REGION Network 14
   RUNG wire#powerrail
      "FC_ANIM_MOTOR"(Input_1 := "MP012-CO", Input_3 := "DB90".Static_6, Input_4 := "MP012-TO", Input_5 := "DB34".Static_24, Output_0 => "DB46".Static_2, Input_0 := wire#w1, Input_2 := wire#w2)
   END_RUNG
   RUNG wire#powerrail
      Contact( "MP012-Marcha" )
      I_Contact( "PRESOSTATO-TORRES" )
   END_RUNG wire#w1
   RUNG wire#powerrail
      Contact( "DB90".Static_110 )
      I_Contact( "DB90".Static_136 )
   END_RUNG wire#w2
   // the same network as SCL:
   "FC_ANIM_MOTOR"(Input_0 := "MP012-Marcha" AND NOT "PRESOSTATO-TORRES",
                   Input_1 := "MP012-CO",
                   Input_2 := "DB90".Static_110 AND NOT "DB90".Static_136,
                   Input_3 := "DB90".Static_6,
                   Input_4 := "MP012-TO",
                   Input_5 := "DB34".Static_24,
                   Output_0 => "DB46".Static_2);
END_REGION

REGION Network 15
   RUNG wire#powerrail
      "FC_ANIM_MOTOR"(Input_1 := "MP013-CO", Input_3 := "DB90".Static_7, Input_4 := "MP013-TO", Input_5 := "DB34".Static_26, Output_0 => "DB46".Static_3, Input_0 := wire#w1, Input_2 := wire#w2)
   END_RUNG
   RUNG wire#powerrail
      Contact( "MP013-Marcha" )
      I_Contact( "PRESOSTATO-TORRES" )
   END_RUNG wire#w1
   RUNG wire#powerrail
      Contact( "DB90".Static_111 )
      I_Contact( "DB90".Static_137 )
   END_RUNG wire#w2
   // the same network as SCL:
   "FC_ANIM_MOTOR"(Input_0 := "MP013-Marcha" AND NOT "PRESOSTATO-TORRES",
                   Input_1 := "MP013-CO",
                   Input_2 := "DB90".Static_111 AND NOT "DB90".Static_137,
                   Input_3 := "DB90".Static_7,
                   Input_4 := "MP013-TO",
                   Input_5 := "DB34".Static_26,
                   Output_0 => "DB46".Static_3);
END_REGION

REGION Network 16
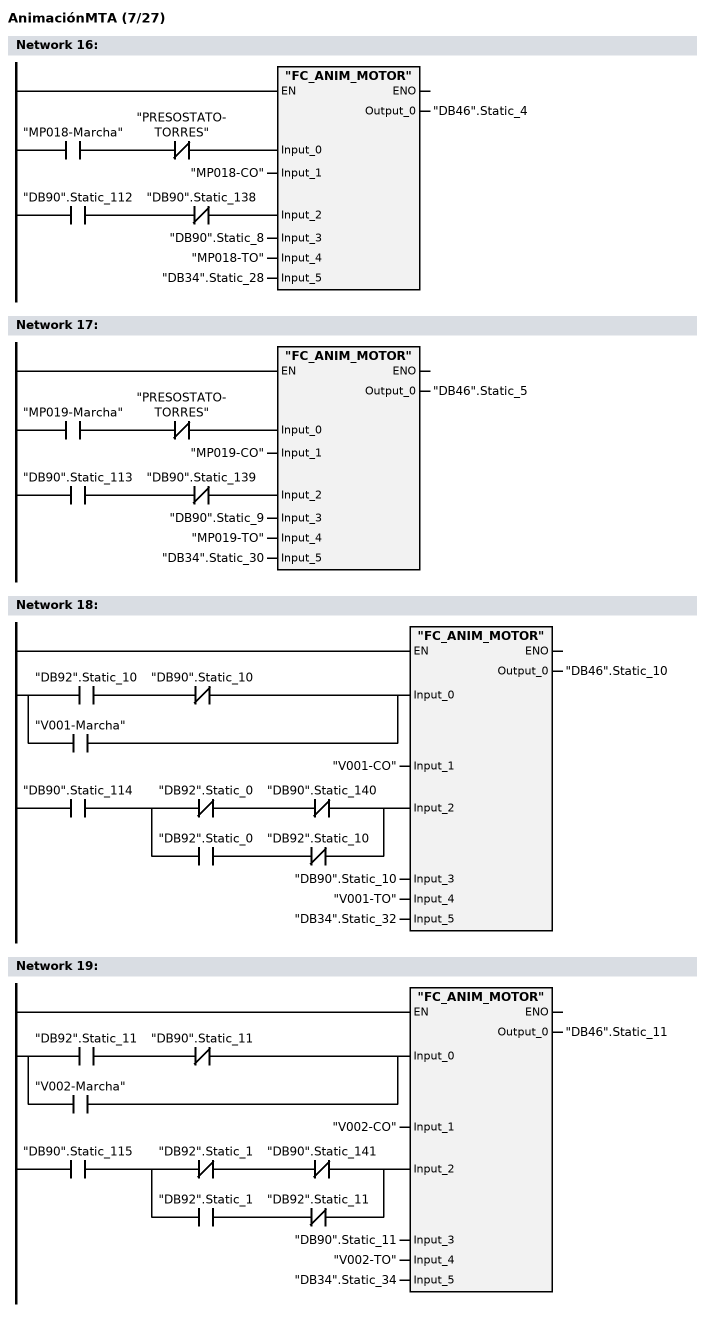
   RUNG wire#powerrail
      "FC_ANIM_MOTOR"(Input_1 := "MP018-CO", Input_3 := "DB90".Static_8, Input_4 := "MP018-TO", Input_5 := "DB34".Static_28, Output_0 => "DB46".Static_4, Input_0 := wire#w1, Input_2 := wire#w2)
   END_RUNG
   RUNG wire#powerrail
      Contact( "MP018-Marcha" )
      I_Contact( "PRESOSTATO-TORRES" )
   END_RUNG wire#w1
   RUNG wire#powerrail
      Contact( "DB90".Static_112 )
      I_Contact( "DB90".Static_138 )
   END_RUNG wire#w2
   // the same network as SCL:
   "FC_ANIM_MOTOR"(Input_0 := "MP018-Marcha" AND NOT "PRESOSTATO-TORRES",
                   Input_1 := "MP018-CO",
                   Input_2 := "DB90".Static_112 AND NOT "DB90".Static_138,
                   Input_3 := "DB90".Static_8,
                   Input_4 := "MP018-TO",
                   Input_5 := "DB34".Static_28,
                   Output_0 => "DB46".Static_4);
END_REGION

REGION Network 17
   RUNG wire#powerrail
      "FC_ANIM_MOTOR"(Input_1 := "MP019-CO", Input_3 := "DB90".Static_9, Input_4 := "MP019-TO", Input_5 := "DB34".Static_30, Output_0 => "DB46".Static_5, Input_0 := wire#w1, Input_2 := wire#w2)
   END_RUNG
   RUNG wire#powerrail
      Contact( "MP019-Marcha" )
      I_Contact( "PRESOSTATO-TORRES" )
   END_RUNG wire#w1
   RUNG wire#powerrail
      Contact( "DB90".Static_113 )
      I_Contact( "DB90".Static_139 )
   END_RUNG wire#w2
   // the same network as SCL:
   "FC_ANIM_MOTOR"(Input_0 := "MP019-Marcha" AND NOT "PRESOSTATO-TORRES",
                   Input_1 := "MP019-CO",
                   Input_2 := "DB90".Static_113 AND NOT "DB90".Static_139,
                   Input_3 := "DB90".Static_9,
                   Input_4 := "MP019-TO",
                   Input_5 := "DB34".Static_30,
                   Output_0 => "DB46".Static_5);
END_REGION

REGION Network 18
   "FC_ANIM_MOTOR"(Input_0 := "V001-Marcha" OR ("DB92".Static_10 AND NOT "DB90".Static_10),
                   Input_1 := "V001-CO",
                   Input_2 := "DB90".Static_114 AND ((NOT "DB92".Static_0 AND NOT "DB90".Static_140) OR ("DB92".Static_0 AND NOT "DB92".Static_10)),
                   Input_3 := "DB90".Static_10,
                   Input_4 := "V001-TO",
                   Input_5 := "DB34".Static_32,
                   Output_0 => "DB46".Static_10);
END_REGION

REGION Network 19
   "FC_ANIM_MOTOR"(Input_0 := "V002-Marcha" OR ("DB92".Static_11 AND NOT "DB90".Static_11),
                   Input_1 := "V002-CO",
                   Input_2 := "DB90".Static_115 AND ((NOT "DB92".Static_1 AND NOT "DB90".Static_141) OR ("DB92".Static_1 AND NOT "DB92".Static_11)),
                   Input_3 := "DB90".Static_11,
                   Input_4 := "V002-TO",
                   Input_5 := "DB34".Static_34,
                   Output_0 => "DB46".Static_11);
END_REGION

REGION Network 20
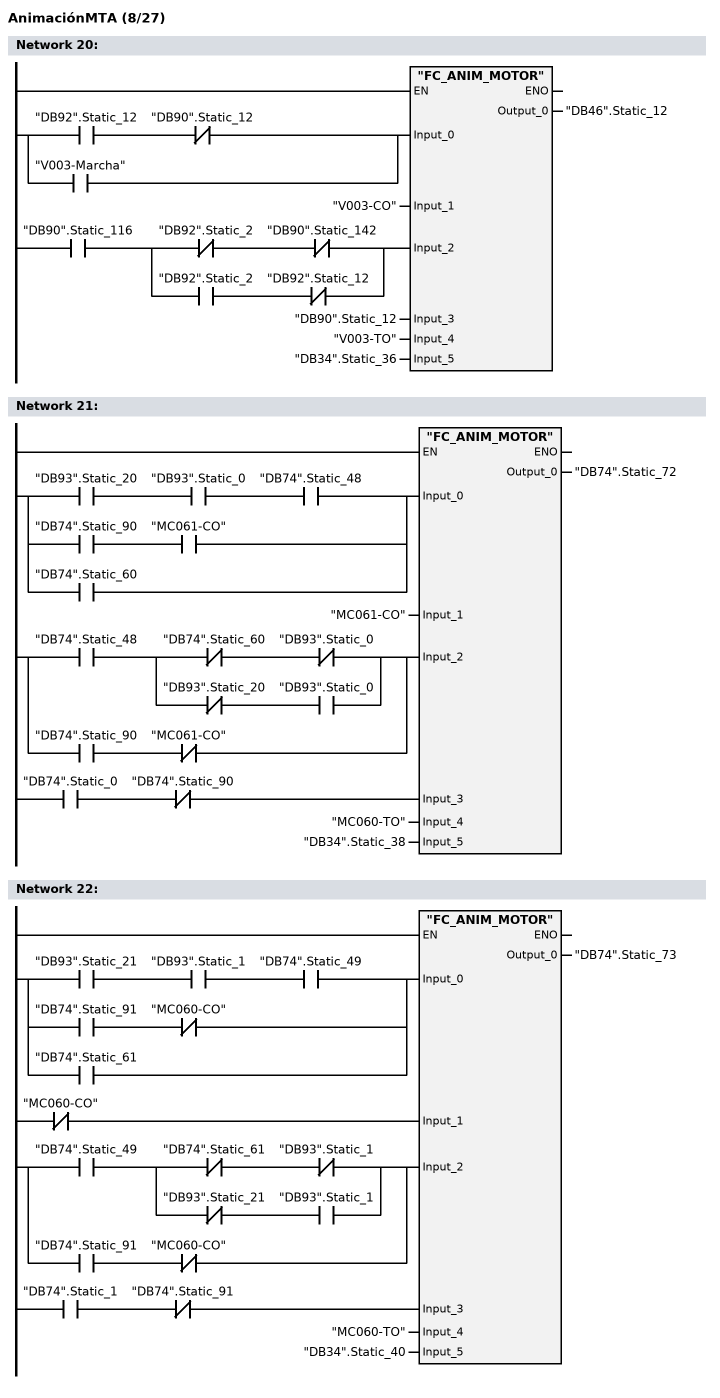
   "FC_ANIM_MOTOR"(Input_0 := "V003-Marcha" OR ("DB92".Static_12 AND NOT "DB90".Static_12),
                   Input_1 := "V003-CO",
                   Input_2 := "DB90".Static_116 AND ((NOT "DB92".Static_2 AND NOT "DB90".Static_142) OR ("DB92".Static_2 AND NOT "DB92".Static_12)),
                   Input_3 := "DB90".Static_12,
                   Input_4 := "V003-TO",
                   Input_5 := "DB34".Static_36,
                   Output_0 => "DB46".Static_12);
END_REGION

REGION Network 21
   "FC_ANIM_MOTOR"(Input_0 := "DB74".Static_60 OR ("DB93".Static_20 AND "DB93".Static_0 AND "DB74".Static_48) OR ("DB74".Static_90 AND "MC061-CO"),
                   Input_1 := "MC061-CO",
                   Input_2 := ("DB74".Static_48 AND ((NOT "DB74".Static_60 AND NOT "DB93".Static_0) OR (NOT "DB93".Static_20 AND "DB93".Static_0))) OR ("DB74".Static_90 AND NOT "MC061-CO"),
                   Input_3 := "DB74".Static_0 AND NOT "DB74".Static_90,
                   Input_4 := "MC060-TO",
                   Input_5 := "DB34".Static_38,
                   Output_0 => "DB74".Static_72);
END_REGION

REGION Network 22
   "FC_ANIM_MOTOR"(Input_0 := "DB74".Static_61 OR ("DB93".Static_21 AND "DB93".Static_1 AND "DB74".Static_49) OR ("DB74".Static_91 AND NOT "MC060-CO"),
                   Input_1 := NOT "MC060-CO",
                   Input_2 := ("DB74".Static_49 AND ((NOT "DB74".Static_61 AND NOT "DB93".Static_1) OR (NOT "DB93".Static_21 AND "DB93".Static_1))) OR ("DB74".Static_91 AND NOT "MC060-CO"),
                   Input_3 := "DB74".Static_1 AND NOT "DB74".Static_91,
                   Input_4 := "MC060-TO",
                   Input_5 := "DB34".Static_40,
                   Output_0 => "DB74".Static_73);
END_REGION

REGION Network 23
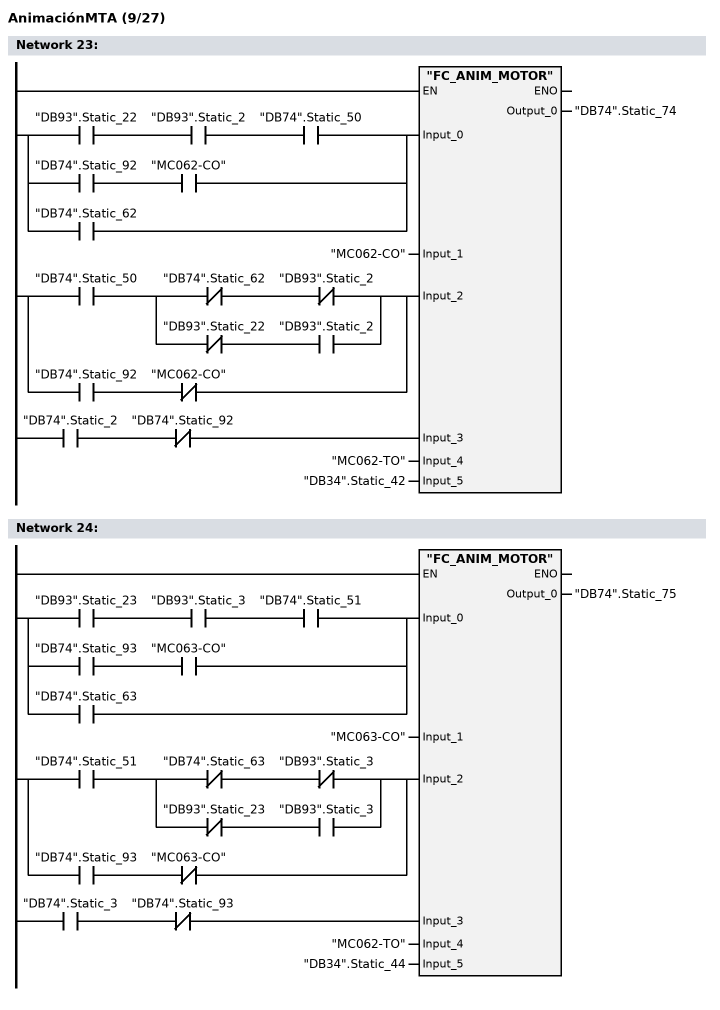
   "FC_ANIM_MOTOR"(Input_0 := "DB74".Static_62 OR ("DB93".Static_22 AND "DB93".Static_2 AND "DB74".Static_50) OR ("DB74".Static_92 AND "MC062-CO"),
                   Input_1 := "MC062-CO",
                   Input_2 := ("DB74".Static_50 AND ((NOT "DB74".Static_62 AND NOT "DB93".Static_2) OR (NOT "DB93".Static_22 AND "DB93".Static_2))) OR ("DB74".Static_92 AND NOT "MC062-CO"),
                   Input_3 := "DB74".Static_2 AND NOT "DB74".Static_92,
                   Input_4 := "MC062-TO",
                   Input_5 := "DB34".Static_42,
                   Output_0 => "DB74".Static_74);
END_REGION

REGION Network 24
   "FC_ANIM_MOTOR"(Input_0 := "DB74".Static_63 OR ("DB93".Static_23 AND "DB93".Static_3 AND "DB74".Static_51) OR ("DB74".Static_93 AND "MC063-CO"),
                   Input_1 := "MC063-CO",
                   Input_2 := ("DB74".Static_51 AND ((NOT "DB74".Static_63 AND NOT "DB93".Static_3) OR (NOT "DB93".Static_23 AND "DB93".Static_3))) OR ("DB74".Static_93 AND NOT "MC063-CO"),
                   Input_3 := "DB74".Static_3 AND NOT "DB74".Static_93,
                   Input_4 := "MC062-TO",
                   Input_5 := "DB34".Static_44,
                   Output_0 => "DB74".Static_75);
END_REGION

REGION Network 25
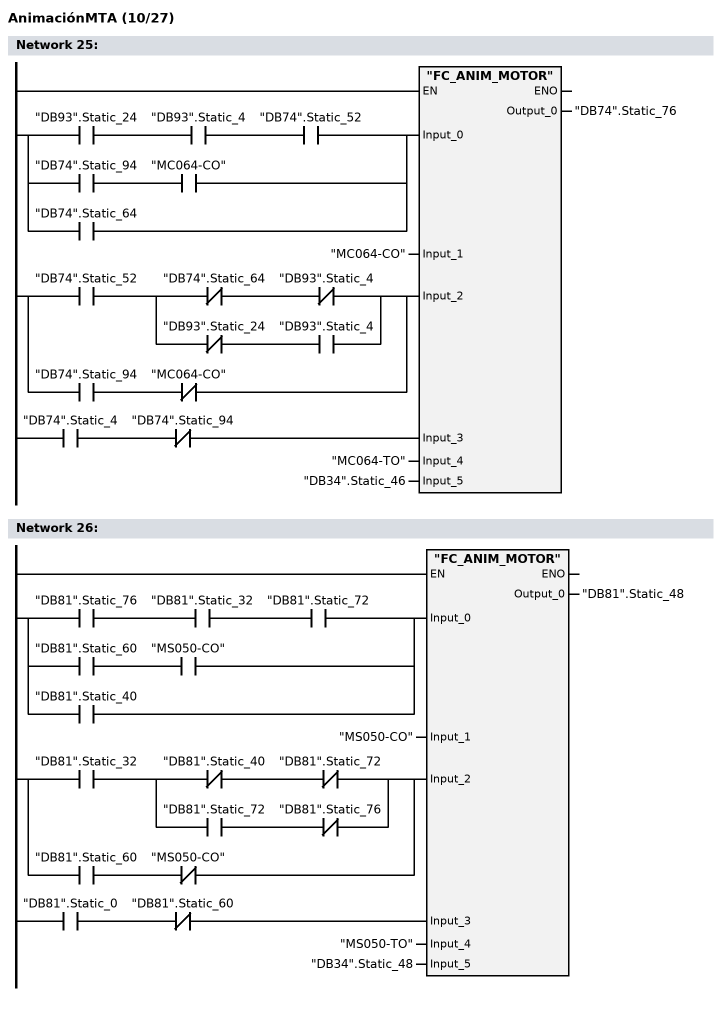
   "FC_ANIM_MOTOR"(Input_0 := "DB74".Static_64 OR ("DB93".Static_24 AND "DB93".Static_4 AND "DB74".Static_52) OR ("DB74".Static_94 AND "MC064-CO"),
                   Input_1 := "MC064-CO",
                   Input_2 := ("DB74".Static_52 AND ((NOT "DB74".Static_64 AND NOT "DB93".Static_4) OR (NOT "DB93".Static_24 AND "DB93".Static_4))) OR ("DB74".Static_94 AND NOT "MC064-CO"),
                   Input_3 := "DB74".Static_4 AND NOT "DB74".Static_94,
                   Input_4 := "MC064-TO",
                   Input_5 := "DB34".Static_46,
                   Output_0 => "DB74".Static_76);
END_REGION

REGION Network 26
   "FC_ANIM_MOTOR"(Input_0 := "DB81".Static_40 OR ("DB81".Static_76 AND "DB81".Static_32 AND "DB81".Static_72) OR ("DB81".Static_60 AND "MS050-CO"),
                   Input_1 := "MS050-CO",
                   Input_2 := ("DB81".Static_32 AND ((NOT "DB81".Static_40 AND NOT "DB81".Static_72) OR ("DB81".Static_72 AND NOT "DB81".Static_76))) OR ("DB81".Static_60 AND NOT "MS050-CO"),
                   Input_3 := "DB81".Static_0 AND NOT "DB81".Static_60,
                   Input_4 := "MS050-TO",
                   Input_5 := "DB34".Static_48,
                   Output_0 => "DB81".Static_48);
END_REGION

REGION Network 27
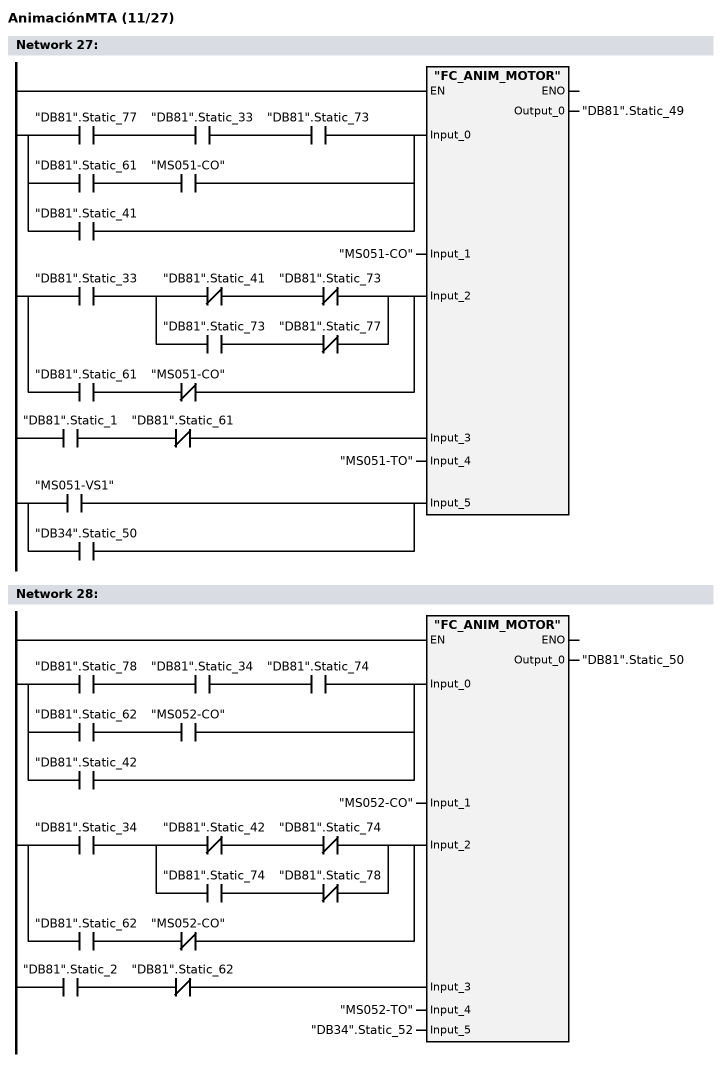
   "FC_ANIM_MOTOR"(Input_0 := "DB81".Static_41 OR ("DB81".Static_77 AND "DB81".Static_33 AND "DB81".Static_73) OR ("DB81".Static_61 AND "MS051-CO"),
                   Input_1 := "MS051-CO",
                   Input_2 := ("DB81".Static_33 AND ((NOT "DB81".Static_41 AND NOT "DB81".Static_73) OR ("DB81".Static_73 AND NOT "DB81".Static_77))) OR ("DB81".Static_61 AND NOT "MS051-CO"),
                   Input_3 := "DB81".Static_1 AND NOT "DB81".Static_61,
                   Input_4 := "MS051-TO",
                   Input_5 := "MS051-VS1" OR "DB34".Static_50,
                   Output_0 => "DB81".Static_49);
END_REGION

REGION Network 28
   "FC_ANIM_MOTOR"(Input_0 := "DB81".Static_42 OR ("DB81".Static_78 AND "DB81".Static_34 AND "DB81".Static_74) OR ("DB81".Static_62 AND "MS052-CO"),
                   Input_1 := "MS052-CO",
                   Input_2 := ("DB81".Static_34 AND ((NOT "DB81".Static_42 AND NOT "DB81".Static_74) OR ("DB81".Static_74 AND NOT "DB81".Static_78))) OR ("DB81".Static_62 AND NOT "MS052-CO"),
                   Input_3 := "DB81".Static_2 AND NOT "DB81".Static_62,
                   Input_4 := "MS052-TO",
                   Input_5 := "DB34".Static_52,
                   Output_0 => "DB81".Static_50);
END_REGION

REGION Network 29
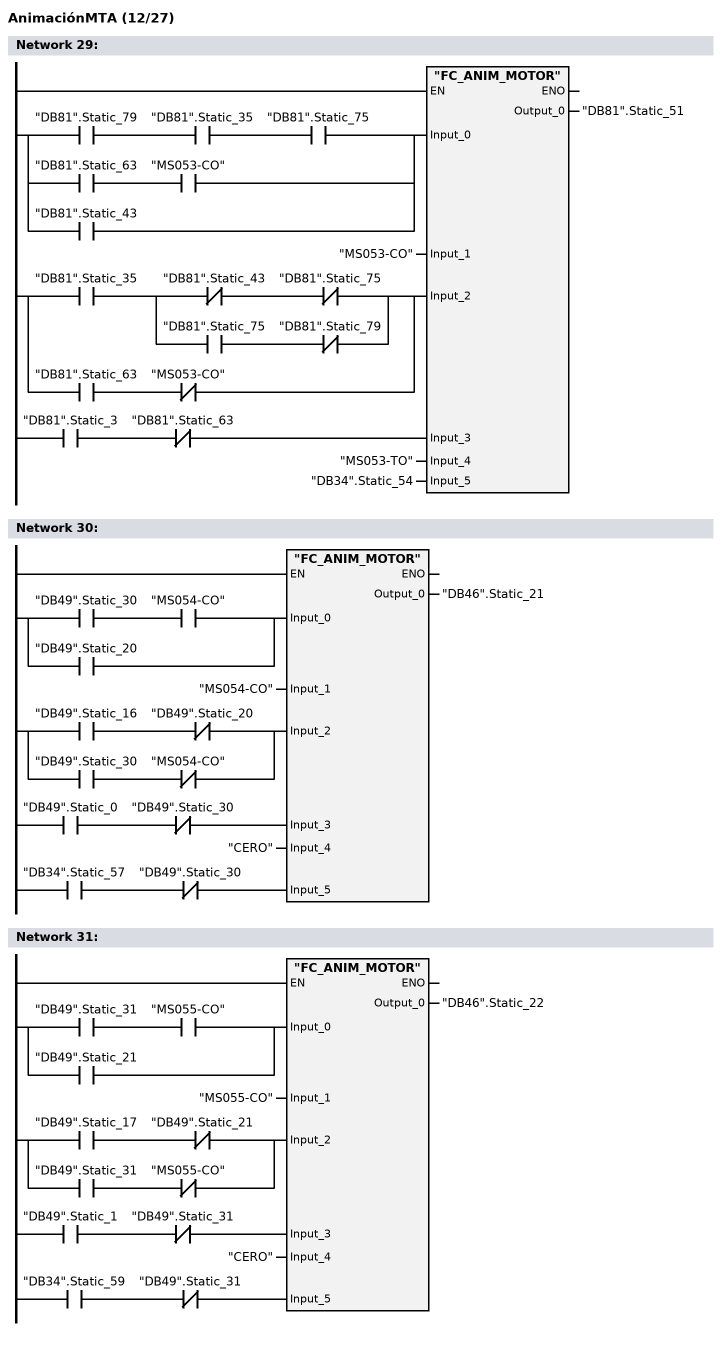
   "FC_ANIM_MOTOR"(Input_0 := "DB81".Static_43 OR ("DB81".Static_79 AND "DB81".Static_35 AND "DB81".Static_75) OR ("DB81".Static_63 AND "MS053-CO"),
                   Input_1 := "MS053-CO",
                   Input_2 := ("DB81".Static_35 AND ((NOT "DB81".Static_43 AND NOT "DB81".Static_75) OR ("DB81".Static_75 AND NOT "DB81".Static_79))) OR ("DB81".Static_63 AND NOT "MS053-CO"),
                   Input_3 := "DB81".Static_3 AND NOT "DB81".Static_63,
                   Input_4 := "MS053-TO",
                   Input_5 := "DB34".Static_54,
                   Output_0 => "DB81".Static_51);
END_REGION

REGION Network 30
   "FC_ANIM_MOTOR"(Input_0 := "DB49".Static_20 OR ("DB49".Static_30 AND "MS054-CO"),
                   Input_1 := "MS054-CO",
                   Input_2 := ("DB49".Static_16 AND NOT "DB49".Static_20) OR ("DB49".Static_30 AND NOT "MS054-CO"),
                   Input_3 := "DB49".Static_0 AND NOT "DB49".Static_30,
                   Input_4 := "CERO",
                   Input_5 := "DB34".Static_57 AND NOT "DB49".Static_30,
                   Output_0 => "DB46".Static_21);
END_REGION

REGION Network 31
   "FC_ANIM_MOTOR"(Input_0 := "DB49".Static_21 OR ("DB49".Static_31 AND "MS055-CO"),
                   Input_1 := "MS055-CO",
                   Input_2 := ("DB49".Static_17 AND NOT "DB49".Static_21) OR ("DB49".Static_31 AND NOT "MS055-CO"),
                   Input_3 := "DB49".Static_1 AND NOT "DB49".Static_31,
                   Input_4 := "CERO",
                   Input_5 := "DB34".Static_59 AND NOT "DB49".Static_31,
                   Output_0 => "DB46".Static_22);
END_REGION

REGION Network 32
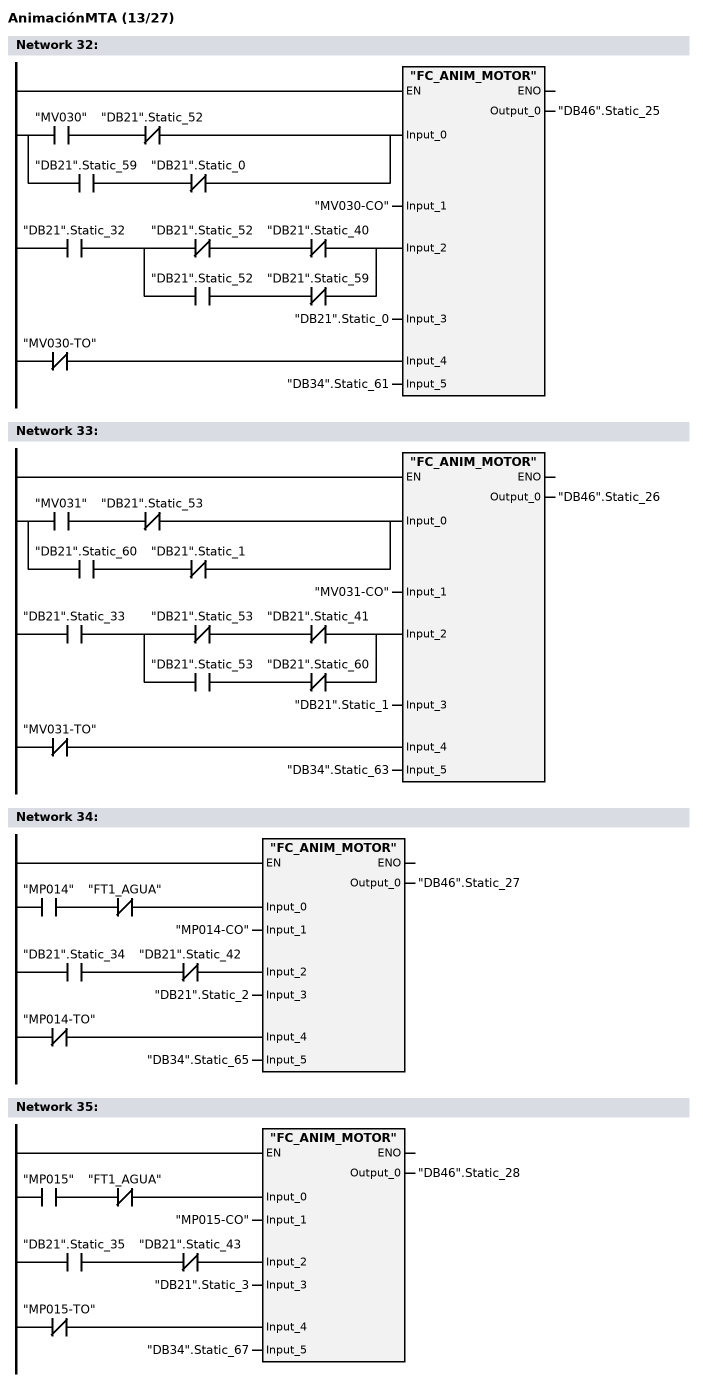
   "FC_ANIM_MOTOR"(Input_0 := ("MV030" AND NOT "DB21".Static_52) OR ("DB21".Static_59 AND NOT "DB21".Static_0),
                   Input_1 := "MV030-CO",
                   Input_2 := "DB21".Static_32 AND ((NOT "DB21".Static_52 AND NOT "DB21".Static_40) OR ("DB21".Static_52 AND NOT "DB21".Static_59)),
                   Input_3 := "DB21".Static_0,
                   Input_4 := NOT "MV030-TO",
                   Input_5 := "DB34".Static_61,
                   Output_0 => "DB46".Static_25);
END_REGION

REGION Network 33
   "FC_ANIM_MOTOR"(Input_0 := ("MV031" AND NOT "DB21".Static_53) OR ("DB21".Static_60 AND NOT "DB21".Static_1),
                   Input_1 := "MV031-CO",
                   Input_2 := "DB21".Static_33 AND ((NOT "DB21".Static_53 AND NOT "DB21".Static_41) OR ("DB21".Static_53 AND NOT "DB21".Static_60)),
                   Input_3 := "DB21".Static_1,
                   Input_4 := NOT "MV031-TO",
                   Input_5 := "DB34".Static_63,
                   Output_0 => "DB46".Static_26);
END_REGION

REGION Network 34
   RUNG wire#powerrail
      "FC_ANIM_MOTOR"(Input_1 := "MP014-CO", Input_3 := "DB21".Static_2, Input_5 := "DB34".Static_65, Output_0 => "DB46".Static_27, Input_0 := wire#w1, Input_2 := wire#w2, Input_4 := wire#w3)
   END_RUNG
   RUNG wire#powerrail
      Contact( "MP014" )
      I_Contact( "FT1_AGUA" )
   END_RUNG wire#w1
   RUNG wire#powerrail
      Contact( "DB21".Static_34 )
      I_Contact( "DB21".Static_42 )
   END_RUNG wire#w2
   RUNG wire#powerrail
      I_Contact( "MP014-TO" )
   END_RUNG wire#w3
   // the same network as SCL:
   "FC_ANIM_MOTOR"(Input_0 := "MP014" AND NOT "FT1_AGUA",
                   Input_1 := "MP014-CO",
                   Input_2 := "DB21".Static_34 AND NOT "DB21".Static_42,
                   Input_3 := "DB21".Static_2,
                   Input_4 := NOT "MP014-TO",
                   Input_5 := "DB34".Static_65,
                   Output_0 => "DB46".Static_27);
END_REGION

REGION Network 35
   RUNG wire#powerrail
      "FC_ANIM_MOTOR"(Input_1 := "MP015-CO", Input_3 := "DB21".Static_3, Input_5 := "DB34".Static_67, Output_0 => "DB46".Static_28, Input_0 := wire#w1, Input_2 := wire#w2, Input_4 := wire#w3)
   END_RUNG
   RUNG wire#powerrail
      Contact( "MP015" )
      I_Contact( "FT1_AGUA" )
   END_RUNG wire#w1
   RUNG wire#powerrail
      Contact( "DB21".Static_35 )
      I_Contact( "DB21".Static_43 )
   END_RUNG wire#w2
   RUNG wire#powerrail
      I_Contact( "MP015-TO" )
   END_RUNG wire#w3
   // the same network as SCL:
   "FC_ANIM_MOTOR"(Input_0 := "MP015" AND NOT "FT1_AGUA",
                   Input_1 := "MP015-CO",
                   Input_2 := "DB21".Static_35 AND NOT "DB21".Static_43,
                   Input_3 := "DB21".Static_3,
                   Input_4 := NOT "MP015-TO",
                   Input_5 := "DB34".Static_67,
                   Output_0 => "DB46".Static_28);
END_REGION

REGION Network 36
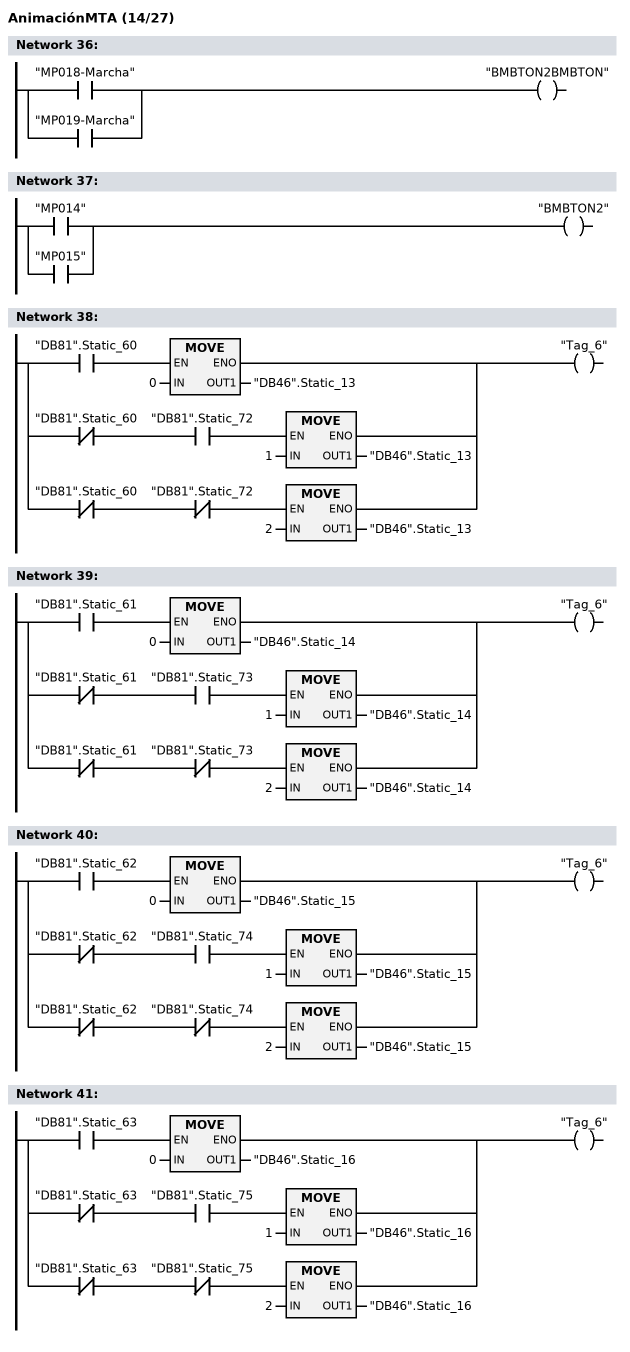
   RUNG wire#powerrail
      Contact( "MP018-Marcha" )
      wire#w1
      Coil( "BMBTON2BMBTON" )
   END_RUNG
   RUNG wire#powerrail
      Contact( "MP019-Marcha" )
   END_RUNG wire#w1
   // the same network as SCL:
   "BMBTON2BMBTON" := "MP018-Marcha" OR "MP019-Marcha";
END_REGION

REGION Network 37
   RUNG wire#powerrail
      Contact( "MP014" )
      wire#w1
      Coil( "BMBTON2" )
   END_RUNG
   RUNG wire#powerrail
      Contact( "MP015" )
   END_RUNG wire#w1
   // the same network as SCL:
   "BMBTON2" := "MP014" OR "MP015";
END_REGION

REGION Network 38
   RUNG wire#powerrail
      Contact( "DB81".Static_60 )
      { S7_GenerateENO := "TRUE" } Move(in := 0, out1 => "DB46".Static_13)
      wire#w1
      Coil( "Tag_6" )
   END_RUNG
   RUNG wire#powerrail
      I_Contact( "DB81".Static_60 )
      Contact( "DB81".Static_72 )
      { S7_GenerateENO := "TRUE" } Move(in := 1, out1 => "DB46".Static_13)
   END_RUNG wire#w1
   RUNG wire#powerrail
      I_Contact( "DB81".Static_60 )
      I_Contact( "DB81".Static_72 )
      { S7_GenerateENO := "TRUE" } Move(in := 2, out1 => "DB46".Static_13)
   END_RUNG wire#w1
   // the same network as SCL:
   // ENO of a box is taken as its EN; it also drops when the box reports an error
   IF "DB81".Static_60 THEN "DB46".Static_13 := 0; END_IF;
   #_w1 := NOT "DB81".Static_60 AND "DB81".Static_72;
   IF #_w1 THEN "DB46".Static_13 := 1; END_IF;
   #_w2 := NOT "DB81".Static_60 AND NOT "DB81".Static_72;
   IF #_w2 THEN "DB46".Static_13 := 2; END_IF;
   "Tag_6" := "DB81".Static_60 OR #_w1 OR #_w2;
END_REGION

REGION Network 39
   RUNG wire#powerrail
      Contact( "DB81".Static_61 )
      { S7_GenerateENO := "TRUE" } Move(in := 0, out1 => "DB46".Static_14)
      wire#w1
      Coil( "Tag_6" )
   END_RUNG
   RUNG wire#powerrail
      I_Contact( "DB81".Static_61 )
      Contact( "DB81".Static_73 )
      { S7_GenerateENO := "TRUE" } Move(in := 1, out1 => "DB46".Static_14)
   END_RUNG wire#w1
   RUNG wire#powerrail
      I_Contact( "DB81".Static_61 )
      I_Contact( "DB81".Static_73 )
      { S7_GenerateENO := "TRUE" } Move(in := 2, out1 => "DB46".Static_14)
   END_RUNG wire#w1
   // the same network as SCL:
   // ENO of a box is taken as its EN; it also drops when the box reports an error
   IF "DB81".Static_61 THEN "DB46".Static_14 := 0; END_IF;
   #_w1 := NOT "DB81".Static_61 AND "DB81".Static_73;
   IF #_w1 THEN "DB46".Static_14 := 1; END_IF;
   #_w2 := NOT "DB81".Static_61 AND NOT "DB81".Static_73;
   IF #_w2 THEN "DB46".Static_14 := 2; END_IF;
   "Tag_6" := "DB81".Static_61 OR #_w1 OR #_w2;
END_REGION

REGION Network 40
   RUNG wire#powerrail
      Contact( "DB81".Static_62 )
      { S7_GenerateENO := "TRUE" } Move(in := 0, out1 => "DB46".Static_15)
      wire#w1
      Coil( "Tag_6" )
   END_RUNG
   RUNG wire#powerrail
      I_Contact( "DB81".Static_62 )
      Contact( "DB81".Static_74 )
      { S7_GenerateENO := "TRUE" } Move(in := 1, out1 => "DB46".Static_15)
   END_RUNG wire#w1
   RUNG wire#powerrail
      I_Contact( "DB81".Static_62 )
      I_Contact( "DB81".Static_74 )
      { S7_GenerateENO := "TRUE" } Move(in := 2, out1 => "DB46".Static_15)
   END_RUNG wire#w1
   // the same network as SCL:
   // ENO of a box is taken as its EN; it also drops when the box reports an error
   IF "DB81".Static_62 THEN "DB46".Static_15 := 0; END_IF;
   #_w1 := NOT "DB81".Static_62 AND "DB81".Static_74;
   IF #_w1 THEN "DB46".Static_15 := 1; END_IF;
   #_w2 := NOT "DB81".Static_62 AND NOT "DB81".Static_74;
   IF #_w2 THEN "DB46".Static_15 := 2; END_IF;
   "Tag_6" := "DB81".Static_62 OR #_w1 OR #_w2;
END_REGION

REGION Network 41
   RUNG wire#powerrail
      Contact( "DB81".Static_63 )
      { S7_GenerateENO := "TRUE" } Move(in := 0, out1 => "DB46".Static_16)
      wire#w1
      Coil( "Tag_6" )
   END_RUNG
   RUNG wire#powerrail
      I_Contact( "DB81".Static_63 )
      Contact( "DB81".Static_75 )
      { S7_GenerateENO := "TRUE" } Move(in := 1, out1 => "DB46".Static_16)
   END_RUNG wire#w1
   RUNG wire#powerrail
      I_Contact( "DB81".Static_63 )
      I_Contact( "DB81".Static_75 )
      { S7_GenerateENO := "TRUE" } Move(in := 2, out1 => "DB46".Static_16)
   END_RUNG wire#w1
   // the same network as SCL:
   // ENO of a box is taken as its EN; it also drops when the box reports an error
   IF "DB81".Static_63 THEN "DB46".Static_16 := 0; END_IF;
   #_w1 := NOT "DB81".Static_63 AND "DB81".Static_75;
   IF #_w1 THEN "DB46".Static_16 := 1; END_IF;
   #_w2 := NOT "DB81".Static_63 AND NOT "DB81".Static_75;
   IF #_w2 THEN "DB46".Static_16 := 2; END_IF;
   "Tag_6" := "DB81".Static_63 OR #_w1 OR #_w2;
END_REGION

REGION Network 42
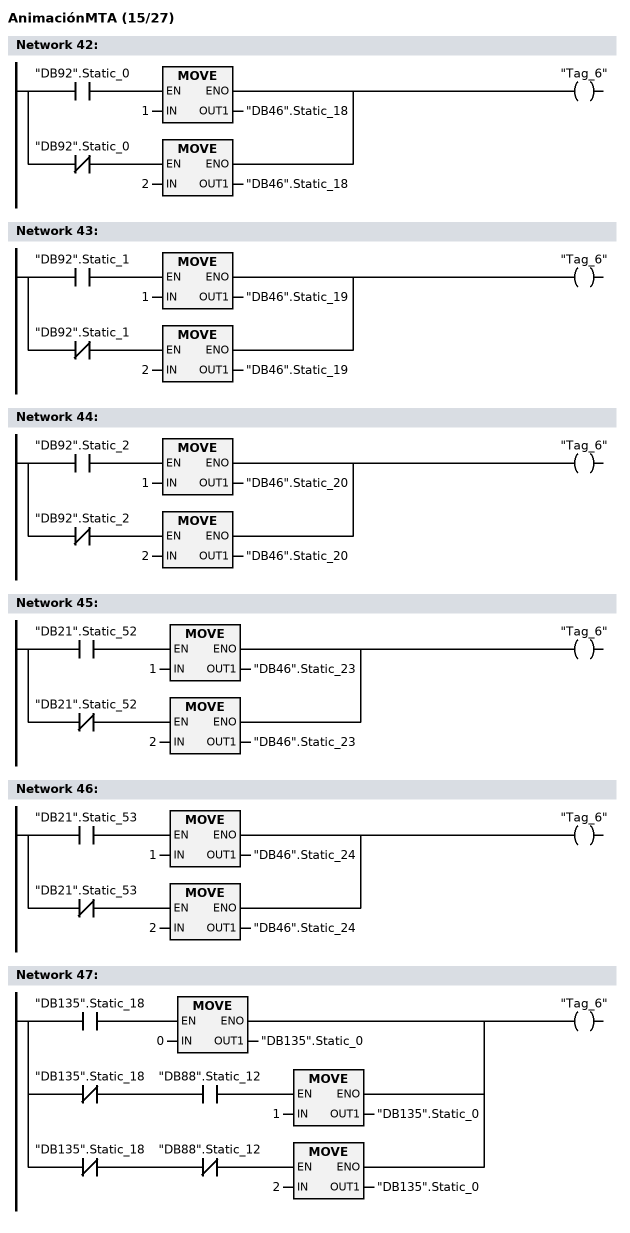
   RUNG wire#powerrail
      Contact( "DB92".Static_0 )
      { S7_GenerateENO := "TRUE" } Move(in := 1, out1 => "DB46".Static_18)
      wire#w1
      Coil( "Tag_6" )
   END_RUNG
   RUNG wire#powerrail
      I_Contact( "DB92".Static_0 )
      { S7_GenerateENO := "TRUE" } Move(in := 2, out1 => "DB46".Static_18)
   END_RUNG wire#w1
   // the same network as SCL:
   // ENO of a box is taken as its EN; it also drops when the box reports an error
   IF "DB92".Static_0 THEN "DB46".Static_18 := 1; END_IF;
   IF NOT "DB92".Static_0 THEN "DB46".Static_18 := 2; END_IF;
   "Tag_6" := "DB92".Static_0 OR NOT "DB92".Static_0;
END_REGION
